
   hm  28. jan.2007   rev 1.1
       modr(x,0) will deliver the result 0

   hm  21. mar 2008    rev 1.2
       use D_trunc for compatibility reasons

   hm  4. apr. 2008    rev 1.3
       added type conversion to avoid warnings under codesys 3.0

   hm  31. oct. 2008   rev 1.4
       changed algorithm to the more common version using floor instead of TRUNC

   hm  10. mar. 2009   rev 1.5
       real constants updated to new systax using dot

   *)
END_FUNCTION

FUNCTION "MUL_ADD" : Real   // FC98, SCL
TITLE = MUL_ADD
{ S7_Optimized_Access := 'FALSE' }
AUTHOR : hugo
FAMILY : MATH
NAME : MUL_ADD
VERSION : 1.1
// this function multiplies an input X with K and adds Offset O to the result.
   VAR_INPUT
      X : Real;
      K : Real;
      O : Real;
   END_VAR
BEGIN


     #MUL_ADD := #X * #K + #O;


   (* revision history
   hm  28. feb 2007
     original version

   hm  11.nov 2007   rev 1.1
     deleted preset values for K and O this makes no sense for a function

   *)
END_FUNCTION

FUNCTION "NEGX" : Real   // FC99, SCL
TITLE = NEGX
{ S7_Optimized_Access := 'FALSE' }
AUTHOR : hugo
FAMILY : MATH
NAME : NEGX
VERSION : 1.0
// This function returns -X
   VAR_INPUT
      X : Real;
   END_VAR
BEGIN


   #NEGX := -#X;

   (* revision history
   hm  26. oct. 2008   rev 1.0
       original version


   *)
END_FUNCTION

FUNCTION "RAD" : Real   // FC100, SCL
TITLE = RAD
{ S7_Optimized_Access := 'FALSE' }
AUTHOR : hugo
FAMILY : MATH
NAME : RAD
VERSION : 1.2
// this function converts Radiant to degrees
// 
// uses: MODR [FC97]
//       FLOOR2 [FC82]
   VAR_INPUT
      deg : Real;
   END_VAR
BEGIN


   #RAD := "MODR"(IN:=0.0174532925199433 * #deg,DIVI:="PI2");

   (*  Enfällt da der Zugriff auf Datenbaustein länger dauert
       RAD := MODR(0.0174532925199433 * DEG, math.PI2);
   *)

   (* revision history
   hm  4. aug 2006     rev 1.0
       original version

   hm  16. oct 2007    rev 1.1
       added modr statement which prohibits rad to become bigger than 2PI

   hm  18. oct 2008    rev 1.2
       using math constants

   *)
END_FUNCTION

FUNCTION "RDM" : Real   // FC101, SCL
TITLE = RDM
{ S7_Optimized_Access := 'FALSE' }
AUTHOR : hugo
FAMILY : MATH
NAME : RDM
VERSION : 1.9
// this function calculates a pseudo random number
// to generate the number it reads the sps timer and calculates a random number between 0 and 1:
// in order to use rdm more then once within one sps cycle it need to be called with different seed numbers LAST.
//  
// uses: T_PLC_MS [FC64]
//       STIME [FB64],IDB_STIME [DB64]
//       BIT_COUNT [FC291]
//       FRACT [FC83]
   VAR_INPUT
      last : Real;
   END_VAR
   VAR_TEMP
      tn : DWord;
      _tn AT tn : Array[0..31] of Bool;
      tc : Int;
   END_VAR
BEGIN


   #tn := "T_PLC_MS"();
   #tc := "BIT_COUNT"(#tn);
   #_tn[7] := #_tn[26];  //tn.31 := tn.2;
   #_tn[6] := #_tn[29];  //tn.30 := tn.5;
   #_tn[5] := #_tn[28];  //tn.29 := tn.4;
   #_tn[4] := #_tn[25];  //tn.28 := tn.1;
   #_tn[3] := #_tn[24];  //tn.27 := tn.0;
   #_tn[2] := #_tn[31];  //tn.26 := tn.7;
   #_tn[1] := #_tn[30];  //tn.25 := tn.6;
   #_tn[0] := #_tn[27];  //tn.24 := tn.3;
   #tn := ROL(IN:=#tn,N:="BIT_COUNT"(#tn)) AND 16#7FFFFFFF OR 16#40000001;  // OR 16#80000001
   #tn := DINT_TO_DWORD(DWORD_TO_DINT(#tn) MOD 71474513 + #tc + 77);
   #RDM := "FRACT"(DINT_TO_REAL(DWORD_TO_DINT(#tn)) / 10000000.0 * ("E"- LIMIT(MN:=0.0,IN:=#last,MX:=1.0)));


   (*
   pt := ADR(temp);
   pt^ := (T_PLC_MS() AND 16#007FFFFF) OR 16#3D000000;
   RDM := fract(modR(temp*e+pi1, PI1-last) + modR(temp*PI1+e + last,e-last));
   *)

   (* revision history
   hm      16. jan 2007        rev 1.0
       original version

   hm      11. nov 2007        rev 1.1
       changed time() into t_plc_ms()

   hm      20. nov 2007        rev 1.2
       changed code of temp calculation to avoid overflow in modr due to resuclt would not fit DINT for high timeer values

   hm      5. jan 2008     rev 1.3
       changed calculation of temp to avoid problem with high values of t_plc_ms

   hm      2. feb 2008     rev 1.4
       changed algorithm to avoind non iec functions and guarantee more randomness

   hm  10. mar. 2008       rev 1.5
       make sure last will be between 0 and 1 to avoid invalid results

   hm  16. mar. 2008       rev 1.6
       added conversion for tc to avoid warnings under codesys 3.0

   hm  18. may. 2008       rev 1.7
       changed constant E to E1

   hm  18. oct. 2008       rev 1.8
       using math constants

   hm  10. mar. 2009       rev 1.9
       real constants updated to new systax using dot

   *)
END_FUNCTION

FUNCTION "RDM2" : Int   // FC102, SCL
TITLE = RDM2
{ S7_Optimized_Access := 'FALSE' }
AUTHOR : hugo
FAMILY : MATH
NAME : RDM2
VERSION : 1.1
// this function calculates an integer pseudo random number
// the random number will be in the range of low <= rdm2 <= high.
// 
// uses: RDM [FC101]
//       T_PLC_MS [FC64] 
//       STIME [FB64],IDB_STIME [DB64] 
//       BIT_COUNT [FC291] 
//       FRACT [FC83]
   VAR_INPUT
      last : Int;
      low : Int;
      high : Int;
   END_VAR
BEGIN


   #RDM2 := REAL_TO_INT(DINT_TO_REAL(TRUNC("RDM"("FRACT"(#last*"PI")) * (#high - #low + 1)) + #low));

   (* revision history
   hm      29. feb 2008        rev 1.0
       original version

   hm      18. oct. 2008       rev 1.1
       using math constants

   *)
END_FUNCTION

FUNCTION "RDMDW" : DWord   // FC103, SCL
TITLE = RDMDW
{ S7_Optimized_Access := 'FALSE' }
AUTHOR : hugo
FAMILY : MATH
NAME : RDMDW
VERSION : 1.2
// this function calculates a DWORD pseudo random number.
// 
// uses: BIT_COUNT [FC291]
//       RDM [FC101]
//       T_PLC_MS [FC64] 
//       STIME [FB64],IDB_STIME [DB64] 
//       FRACT [FC83]
   VAR_INPUT
      last : DWord;
   END_VAR
   VAR_TEMP
      RX : Real;
      "M" : Real;
   END_VAR
BEGIN


   #"M" := "BIT_COUNT"(#last);
   #RX := "RDM"("FRACT"(#"M"*"PI"));
   #RDMDW := SHL(IN:=DINT_TO_DWORD(REAL_TO_DINT(#RX*65535)),N:=16);
   #RX := "RDM"("FRACT"(#"M" * "E"));
   #RDMDW := #RDMDW OR (DINT_TO_DWORD(REAL_TO_DINT(#RX*65535)) AND 16#0000FFFF);

   (* revision history
   hm      14. mar 2008        rev 1.0
       original version

   hm      18. may. 2008       rev 1.1
       changed constant E to E1

   hm      18. oct. 2008       rev 1.2
       using math constants

   *)
END_FUNCTION

FUNCTION "RND" : Real   // FC104, SCL
TITLE = RND
{ S7_Optimized_Access := 'FALSE' }
AUTHOR : hugo
FAMILY : MATH
NAME : RND
VERSION : 1.2
// this function rounds a real down to n digits total.
// round(3.1415,2) = 3.1
// 
// uses: EXPN [FC78]
//       CEIL [FC66]
   VAR_INPUT
      X : Real;
      N : Int;
   END_VAR
   VAR_TEMP
      "M" : Real;
   END_VAR
BEGIN


   IF #X = 0.0 THEN
       #RND := 0.0;
   ELSE
       #"M" := "EXPN"(X:=10.0, N:=#N - "CEIL"((LN(ABS(#X))/LN(10))));
       #RND := DINT_TO_REAL(REAL_TO_DINT(#X * #"M")) / #"M";
   END_IF;


   (* revision history
   hm  11. mar 2008    rev 1.0
       original version

   hm  26. oct. 2008   rev 1.1
       code optimization

   hm  10. mar. 2009   rev 1.2
       real constants updated to new systax using dot

   *)
END_FUNCTION

FUNCTION "ROUND" : Real   // FC105, SCL
TITLE = ROUND
{ S7_Optimized_Access := 'FALSE' }
AUTHOR : hugo
FAMILY : MATH
NAME : ROUND
VERSION : 1.5
// this function rounds a real down to n digits behind the comma.
// round(3.1415,1) = 3.1
   VAR_INPUT
      in : Real;
      N : Int;
   END_VAR
   VAR_TEMP
      X : Real;
   END_VAR
BEGIN


   //x := setup.DECADES[LIMIT(0,n,8)];
   CASE LIMIT(MN:=0, IN:=#N, MX:=8) OF
       1 :           #X:= 10;
       2 :           #X:= 100;
       3 :           #X:= 1000;
       4 :           #X:= 10000;
       5 :           #X:= 100000;
       6 :           #X:= 1000000;
       7 :           #X:= 10000000;
       8 :           #X:= 100000000;
   ELSE: 
       #X:= 1;
   END_CASE ;

   #ROUND := DINT_TO_REAL(REAL_TO_DINT(#in * #X)) / #X;


   (* revision history
   hm  1. sep 2006 rev 1.0
       original version

   hm  2. dec 2007 rev 1.1
       changed code for better performance

   hm  8. jan 2008 rev 1.2
       further improvement in performance

   hm 11. mar. 2008    rev 1.3
       corrected an error with negative numbers
       use real_to_dint instead of trunc

   hm  16. mar 2008    rev 1.4
       added type conversion to avoid warning under codesys 3.0

   hm  25. oct. 2008   rev 1.5
       new code using global constants decades
   *)
END_FUNCTION

FUNCTION "SGN" : Int   // FC106, SCL
TITLE = SGN
{ S7_Optimized_Access := 'FALSE' }
AUTHOR : hugo
FAMILY : MATH
NAME : SGN
VERSION : 1.1
// sgn returns 0 when X = 0 , -1 when X < 1 and +1 when X > 1
   VAR_INPUT
      X : Real;
   END_VAR
BEGIN


     IF #X > 0.0 THEN
       #SGN := 1;
     ELSIF #X < 0.0 THEN
       #SGN := -1;
     ELSE
       #SGN := 0;
     END_IF;

   (* revision histroy
   hm  16. oct 2007  rev 1.0
     original version

   hm  11. nov 2007  rev 1.1
     changed type of function from real to int
   *)
END_FUNCTION

FUNCTION "SIGMOID" : Real   // FC107, SCL
TITLE = SIGMOID
{ S7_Optimized_Access := 'FALSE' }
AUTHOR : hugo
FAMILY : MATH
NAME : SIGMOID
VERSION : 1.2
// this function calculates the sigmoid function
   VAR_INPUT
      X : Real;
   END_VAR
BEGIN


   IF #X > 20.0 THEN
       #SIGMOID := 1.0;
   ELSIF #X < -85.0 THEN
       #SIGMOID := 0.0;
   ELSE
       #SIGMOID := 1.0 / (1.0 + EXP(-#X));
   END_IF;


   (* revision history
   hm  10.12.2007      rev 1.0
       original version

   hm    11. mar. 2008       rev 1.1
       extended range of valid inputs to +inv / -inv

   hm 10. mar. 2009        rev 1.2
       real constants updated to new systax using dot

   *)
END_FUNCTION

FUNCTION "SIGN_I" : Bool   // FC108, SCL
TITLE = SIGN_I
{ S7_Optimized_Access := 'FALSE' }
AUTHOR : hugo
FAMILY : MATH
NAME : SIGN_I
VERSION : 1.3
// this function return true if the integer input is negative
   VAR_INPUT
      IN : DInt;
   END_VAR
BEGIN


   #SIGN_I := #IN < 0;

   (* revision history
   hm 3.3.2007 rev 1.1
       changed method of function for better compatibility to other systems

   hm  1.12.2007   rev 1.2
       changed code to improve performance

   hm  27. oct. 2008   rev 1.3
       changed type of input to dint
   *)
END_FUNCTION

FUNCTION "SIGN_R" : Bool   // FC109, SCL
TITLE = SIGN_R
{ S7_Optimized_Access := 'FALSE' }
AUTHOR : hugo
FAMILY : MATH
NAME : SIGN_R
VERSION : 1.4
// this function return true if the real input is negative
   VAR_INPUT
      in : Real;
   END_VAR
BEGIN


   #SIGN_R := #in < 0.0;


   (* revision history
   hm 19.1.2007    rev 1.1
       changed method of function for better compatibility to other systems

   hm  1.12.2007   rev 1.2
       changed code to improve performance

   hm  14. jun. 2008   rev 1.3
       improved performace

   hm 10. mar. 2009    rev 1.4
       real constants updated to new systax using dot
   *)
END_FUNCTION

FUNCTION "SINC" : Real   // FC110, SCL
TITLE = SINC
{ S7_Optimized_Access := 'FALSE' }
AUTHOR : hugo
FAMILY : MATH
NAME : SINC
VERSION : 1.2
// this function calculates the sinc function.
   VAR_INPUT
      X : Real;
   END_VAR
BEGIN


   IF #X = 0.0 THEN
       #SINC := 1.0;
   ELSE
       #SINC := SIN(#X) / #X;
   END_IF;


   (* revision histroy
   hm  11. mar. 2008   rev 1.0
       original version

   hm  1.12.2007   rev 1.1
       changed code to improove performance

   hm 10. mar. 2009    rev 1.2
       real constants updated to new systax using dot

   *)
END_FUNCTION

FUNCTION "SINH" : Real   // FC111, SCL
TITLE = SINH
{ S7_Optimized_Access := 'FALSE' }
AUTHOR : hugo
FAMILY : MATH
NAME : SINH
VERSION : 1.3
// this function calculates the sin hyperbolicus
   VAR_INPUT
      X : Real;
   END_VAR
BEGIN


   IF ABS(#X) < 2.0E-3 THEN
       #SINH := #X;
   ELSE
       #SINH := (EXP(#X) - EXP(-#X)) * 0.5;
   END_IF;

   (* revision history
   hm  12.1.2007   rev 1.0
       original version

   hm  1.12.2007   rev 1.1
       changed code to improve performance

   hm  5. jan 2008 rev 1.2
       further performance improvement

   hm  11. mar 2008    rev 1.3
       improved accuracy around 0

   *)
END_FUNCTION

FUNCTION "SQRTN" : Real   // FC112, SCL
TITLE = SQRTN
{ S7_Optimized_Access := 'FALSE' }
AUTHOR : hugo
FAMILY : MATH
NAME : SQRTN
VERSION : 1.3
// this function calculates the nth root function of X according to the formula sqrtn = x^(1/n).
   VAR_INPUT
      X : Real;
      N : Int;
   END_VAR
BEGIN


   IF #N > 0 THEN
       #SQRTN := EXP(LN(#X) / INT_TO_REAL(#N));
   ELSE
       #SQRTN := 0.0;
   END_IF;


   (* revision history
   hm      12 jan 2007 rev 1.0
       original version

   hm      2. dec 2007 rev 1.1
       changed code for better performance

   hm      11. mar 2008    rev 1.2
       added result 0 for compatibility reasons

   hm 10. mar. 2009    rev 1.3
       added type conversions for compatibility reasons

   *)
END_FUNCTION

FUNCTION "TANC" : Real   // FC113, SCL
TITLE = TANC
{ S7_Optimized_Access := 'FALSE' }
AUTHOR : hugo
FAMILY : MATH
NAME : TANC
VERSION : 1.1
// this function calculates the tanc function.
   VAR_INPUT
      X : Real;
   END_VAR
BEGIN


   IF #X = 0.0 THEN
       #TANC := 1.0;
   ELSE
       #TANC := TAN(#X) / #X;
   END_IF;


   (* revision histroy
   hm  23. oct. 2008   rev 1.0
       original version

   hm 10. mar. 2009    rev 1.1
       real constants updated to new systax using dot

   *)
END_FUNCTION

FUNCTION "TANH" : Real   // FC114, SCL
TITLE = TANH
{ S7_Optimized_Access := 'FALSE' }
AUTHOR : hugo
FAMILY : MATH
NAME : TANH
VERSION : 1.3
// this function calculates the tangens hyperbolicus
   VAR_INPUT
      X : Real;
   END_VAR
BEGIN


   IF #X > 20.0 THEN
       #TANH := 1.0;
   ELSIF #X < -20.0 THEN
       #TANH := -1.0;
   ELSE
       #TANH := 1.0 - 2.0 / (EXP(2.0 * #X) + 1.0);
   END_IF;


   (* revision hisdtory
   hm      12.1.2007       rev 1.0
       original version

   hm      1.12.2007       rev 1.1
       changed code to improve performance

   hm      10. mar 2008    rev 1.2
       corrected an error in formula
       extended range of valid inputs to +/- INV

   hm 10. mar. 2009    rev 1.3
       real constants updated to new systax using dot

   *)
END_FUNCTION

FUNCTION "WINDOW" : Bool   // FC115, SCL
TITLE = WINDOW
{ S7_Optimized_Access := 'FALSE' }
AUTHOR : hugo
FAMILY : MATH
NAME : WINDOW
VERSION : 1.1
// this checks a signal if the signal is between the upper and lower limit
   VAR_INPUT
      low : Real;
      in : Real;
      high : Real;
   END_VAR
BEGIN


   #WINDOW := #in < #high AND #in > #low;


   (* revision history
   hm  22.1.2007   rev 1.1
       changed the order of inputs to low, in, high

   *)
END_FUNCTION

FUNCTION "WINDOW2" : Bool   // FC116, SCL
TITLE = WINDOW2
{ S7_Optimized_Access := 'FALSE' }
AUTHOR : hugo
FAMILY : MATH
NAME : WINDOW2
VERSION : 1.0
// this checks a signal if the signal is between the upper and lower limit including the two limits
   VAR_INPUT
      low : Real;
      in : Real;
      high : Real;
   END_VAR
BEGIN


   #WINDOW2 := #in <= #high AND #in >= #low;


   (* revision history
   hm  31.10.2007  rev 1.0
     original version

   *)
END_FUNCTION

FUNCTION "BIT_COUNT" : Int   // FC291, SCL
TITLE = BIT_COUNT
{ S7_Optimized_Access := 'FALSE' }
AUTHOR : hugo
FAMILY : GATE
NAME : BITCT
VERSION : 1.1
// BIT_COUNT counts the amount True of bits in a dword.
// for exabple: bit_count(3) returns 2 because two bits (bits 0 and 1) are true and all others are false.
   VAR_INPUT
      IN : DWord;
   END_VAR
   VAR_TEMP
      temp : DWord;
      attemp AT temp : Array[0..31] of Bool;
   END_VAR
BEGIN


     #BIT_COUNT := 0;
     #temp := #IN;

     WHILE DWORD_TO_DINT(#temp) <> 0 DO
       IF #attemp[24] THEN #BIT_COUNT := #BIT_COUNT +1; END_IF;
       #temp := SHR(IN:=#temp,N:=1);
     END_WHILE;

   (* revision history
   5.7.2007  rev 1.0    original version

   10.9.2007  rev 1.1    hm
     changed algorithm for better performace
     the execution time has reduced by a factor of 5
     deleted unused variable temp
   *)
END_FUNCTION

FUNCTION "LAMBERT_W" : Real   // FC414, SCL
TITLE = LAMBERT_W
{ S7_Optimized_Access := 'FALSE' }
AUTHOR : hugo
FAMILY : MATH
NAME : LAMBERT
VERSION : 1.1
// this function calculates the lambert_w function.
   VAR_INPUT
      X : Real;
   END_VAR
   VAR_TEMP
      w : Real;
      i : Int;
      we : Real;
      w1e : Real;
      last : DWord;
      ewx : Real;
   END_VAR
BEGIN


   (* check for valid input and return -1000 if too low *)
   IF #X < -0.367879441171442 THEN
       #LAMBERT_W := -1000.0;
       RETURN;
   (* return 0 if x = 0 *)
   ELSIF #X = 0.0 THEN
       RETURN;
   (* first an estimate is calculated *)
   ELSIF #X <= 500.0 THEN
       #w := LN(#X + 1.0);
       #w := 0.665 * (1.0 + 0.0195 * #w) * #w + 0.04;
   ELSE
       #w := LN(#X - 4.0) - (1.0 - 1.0/LN(#X)) * LN(LN(#X));
   END_IF;
   (* use estimate to calculate exact result *)
   FOR #i := 0 TO 5 DO
       #ewx := EXP(#w);
       #we := #w * #ewx - #X;
       #w1e := (#w + 1.0) * #ewx;
       #last := REAL_TO_DWORD(#w) AND 16#FFFF_FFFC;
       #w := #w - (#we / (#w1e - (#w+2.0) * #we / (2.0 * #w + 2.0)));
       IF (REAL_TO_DWORD(#w) AND 16#FFFF_FFFC) = #last THEN EXIT; END_IF;
   END_FOR;
   #LAMBERT_W := #w;


   (* revision hisdtory
   hm  26. oct. 2008   rev 1.0
       original version

   hm  10. mar. 2009   rev 1.1
       real constants updated to new systax using dot

   *)
END_FUNCTION

FUNCTION "REAL_TO_FRAC" : "FRACTION"   // FC427, SCL
TITLE = REAL_TO_FRAC
{ S7_Optimized_Access := 'FALSE' }
AUTHOR : alex
FAMILY : MATH
NAME : R2FRAC
VERSION : 1.0
// this function calculates the closest fraction for a real number
// 
// uses: FRACTION [UDT19]
   VAR_INPUT
      X : Real;
      N : Int;
   END_VAR
   VAR_TEMP
      temp : DInt;
      sign : Bool;
      X_gerundet : DInt;
      X_ohne_Nachkomma : Real;
      Numerator : DInt;
      Denominator : DInt;
      Numerator_old : DInt;
      Denominator_old : DInt;
      tX : Real;
      tREAL_TO_FRAC : "FRACTION";
   END_VAR
BEGIN


   #Numerator := 1; (* Initialwert Zaehler  *)
   #Denominator := 0; (* Initialwert Nenner *)
   #Numerator_old := 0; (* Initialwert Zaehler der letzten Berechnung  *)
   #Denominator_old := 1; (* Initialwert Zaehler der letzten Berechnung   *)
   #tX := #X;

   (*
   numerator := 1;                     (* Zaehler Initialwert *)
   denominator := 0;                   (* Nenner  Initialwert *)
   numerator_old := 0;
   denominator_old :=1;
   *)

   IF #tX < 0.0 THEN
     #sign := TRUE;               (* Vorzeichen merken *)
     #tX := ABS(#tX);              (* Absolutwert berechnen *)
   END_IF;

   (*
   sign := SIGN_R(X);                    
   X := ABS(X);                      
   *)

   REPEAT
     #X_gerundet := REAL_TO_DINT(#tX);

     (* Zaehler berechnen *)
     #temp := #Numerator * #X_gerundet + #Numerator_old;   (* Zaehler um Vorkammawert erweitern *)
     #Numerator_old := #Numerator;             (* Zaehler der letzten Berechnung speichern *)
     #Numerator := #temp;                  (* Zaehler dieser Berechnung speichern *)

     (* Nenner berechnen *)
     #temp := #Denominator * #X_gerundet + #Denominator_old; (* Nenner um Vorkammawert erweitern *)
     #Denominator_old := #Denominator;           (* Nenner der letzten Berechnung speichern *)
     #Denominator := #temp;                (* Nenner dieser Berechnung speichern *)

     (* Restwert berechnen *)
     #X_ohne_Nachkomma := DINT_TO_REAL(#X_gerundet);
     IF #tX = #X_ohne_Nachkomma THEN            (* Bruch geht ohne Rest auf *)
       IF ABS(#Denominator) <= #N THEN         (* kein Rundungsfehler *)
         #Numerator_old := #Numerator;         (* Numerator_old wird von Funktion zurückgegeben *)
         #Denominator_old := #Denominator;       (* Denominator_old wird von Funktion zurückgegeben *)
       END_IF;
       EXIT;                     (* keine weitere Berechnung notwendig *)
     ELSE
       #tX := 1.0 / (#tX - #X_ohne_Nachkomma);        (* Kehrwert vom Rest -> Neuer Bruch *)
     END_IF;

   UNTIL
     ( ABS(#Denominator) > #N )
   END_REPEAT;

   (* correct sign if X was negative *)
   IF #sign THEN
     #tREAL_TO_FRAC.NUMERATOR := -1 * ABS(DINT_TO_INT(#Numerator_old));
   ELSE
     #tREAL_TO_FRAC.NUMERATOR :=  ABS(DINT_TO_INT(#Numerator_old));
   END_IF;

   #tREAL_TO_FRAC.DENOMINATOR := ABS(DINT_TO_INT(#Denominator_old));

   #REAL_TO_FRAC := #tREAL_TO_FRAC;


   (* revision history
   hm    19. jan. 2011 rev 1.0
     original version

   ad    06. apr. 2011 rev 1.1
     optimized code
   *)
END_FUNCTION

FUNCTION "GCD" : Int   // FC431, SCL
TITLE = GCD
{ S7_Optimized_Access := 'FALSE' }
AUTHOR : hugo
FAMILY : MATH
NAME : GCD
VERSION : 1.0
// this function calculates the gretaest common divisor of two numbers A and B
   VAR_INPUT
      "A" : DInt;
      "B" : DInt;
   END_VAR
   VAR_TEMP
      t : DInt;
      tA : DInt;
      _A AT tA : Array[0..31] of Bool;
      tB : DInt;
      _B AT tB : Array[0..31] of Bool;
   END_VAR
BEGIN


   #tA := #"A";
   #tB := #"B";

   IF #tA = 0 THEN
     #GCD := DINT_TO_INT(ABS(#tB));
   ELSIF #tB = 0 THEN
     #GCD := DINT_TO_INT(ABS(#tA));
   ELSE
     #tA := ABS(#tA);
     #tB := ABS(#tB);
     #GCD := 1;
     WHILE NOT(#_A[24] OR #_B[24]) DO
       #tA := DWORD_TO_DINT(SHR(IN:=DINT_TO_DWORD(#tA),N:=1));
       #tB := DWORD_TO_DINT(SHR(IN:=DINT_TO_DWORD(#tB),N:=1));
       #GCD := WORD_TO_INT(SHL(IN:=INT_TO_WORD(#GCD),N:=1));
     END_WHILE;
     WHILE #tA > 0 DO
       IF NOT(#_A[24]) THEN #tA := DWORD_TO_DINT(SHR(IN:=DINT_TO_DWORD(#tA),N:=1));
       ELSIF NOT(#_B[24]) THEN #tB := DWORD_TO_DINT(SHR(IN:=DINT_TO_DWORD(#tB),N:=1));
       ELSE
         #t:= DWORD_TO_DINT(SHR(IN:=DINT_TO_DWORD(ABS(#tA-#tB)),N:=1));
         IF #tA < #tB THEN #tB := #t; ELSE #tA := #t; END_IF;
       END_IF;
     END_WHILE;
     #GCD := #GCD * DINT_TO_INT(#tB);
   END_IF;


   (* revision history
   hm  19. jan. 2011 rev 1.0
     original version

   *)
END_FUNCTION

// ===== PLC "Mathematical Array"  Unspecific CPU S7 300 =====

VAR_GLOBAL CONSTANT   // PLC tag table "STEP7 classic symbols"
   "debug" : Bool := FALSE;
   "N" : Int := 0;
   "offset" : Int := 0;
   "E" : Real := 2.71828182845904523536028747135266249;   // Eulersche Konstante
   "PI" : Real := 3.14159265358979323846264338327950288;
   "offset_1" : DWord := 0;
END_VAR

DATA_BLOCK "IDB_STIME"   // DB64
{ S7_Optimized_Access := 'FALSE' }
AUTHOR : dalbi
FAMILY : MEASURE
VERSION : 0.0
// stored: InstanceOfName STIME
"STIME"
BEGIN
END_DATA_BLOCK

FUNCTION_BLOCK "_ARRAY_ABS"   // FB5, SCL
TITLE = _ARRAY_ABS
{ S7_Optimized_Access := 'FALSE' }
AUTHOR : hugo
FAMILY : ARFUNCT
NAME : AR_ABS
VERSION : 1.0
// this function will calculate the absolute value of each element of the array and stroe the result instead of the element.
// Array[i] := ABS(ARRAY[i]).
// the function needs to be called:    array_avg(adr("array"),sizeof("array"));
// because this function works with pointers its very time efficient and it needs no extra memory.
   VAR_INPUT
      pt : Pointer;
      _pt AT pt : Struct
         DBNr : Word;
         Adr : DWord;
      END_STRUCT;
      size : Int;
   END_VAR
   VAR_OUTPUT
      _ABS : Bool;
   END_VAR
   VAR_TEMP
      i : Int;
      stop : Int;
      Adr : Int;
      DB_LENGTH : Word;
      WRITE_PROT : Bool;
      rTEST_DB : Int;
   END_VAR
BEGIN


   #_ABS := FALSE;

   (* test data block *)
   #rTEST_DB := TEST_DB(DB_NUMBER := #_pt.DBNr ,DB_LENGTH => #DB_LENGTH ,WRITE_PROT => #WRITE_PROT);
   (* End if TEST_DB <> 0 = Error *)
   IF #rTEST_DB <> 0 THEN RETURN; END_IF;
   (* End if data block to short *) 
   IF WORD_TO_INT(#DB_LENGTH)/4 < #size THEN RETURN; END_IF;
   (* calculate adress for first data *)  
   #Adr := DWORD_TO_INT(SHR(IN:=SHL(IN:=#_pt.Adr,N:=8),N:=11));

   (* code *)
   #stop := #size - 1;   //stop := SHR(size,2)-1;
   FOR #i := 0 TO #stop DO
       WORD_TO_BLOCK_DB(#_pt.DBNr).DD(#Adr+#i*4) := REAL_TO_DWORD(ABS(DWORD_TO_REAL(WORD_TO_BLOCK_DB(#_pt.DBNr).DD(#Adr+#i*4))));
   END_FOR;

   #_ABS := TRUE;


   (* revision history
   hm  2. apr 2008     rev 1.0
       original version

   *)
END_FUNCTION_BLOCK

FUNCTION_BLOCK "_ARRAY_ADD"   // FB6, SCL
TITLE = _ARRAY_ADD
{ S7_Optimized_Access := 'FALSE' }
AUTHOR : hugo
FAMILY : ARFUNCT
NAME : AR_ADD
VERSION : 1.0
// this function will add an offset X to each element of the array and stroe the result instead of the element.
// Array[i] := ARRAY[i] + X.
// the function needs to be called:    array_avg(adr("array"),sizeof("array"));
// because this function works with pointers its very time efficient and it needs no extra memory.
   VAR_INPUT
      pt : Pointer;
      _pt AT pt : Struct
         DBNr : Word;
         Adr : DWord;
      END_STRUCT;
      size : Int;
      X : Real;
   END_VAR
   VAR_OUTPUT
      _ADD : Bool;
   END_VAR
   VAR_TEMP
      i : Int;
      stop : Int;
      Adr : Int;
      DB_LENGTH : Word;
      WRITE_PROT : Bool;
      rTEST_DB : Int;
   END_VAR
BEGIN


   #_ADD := FALSE;

   (* test data block *)
   #rTEST_DB := TEST_DB(DB_NUMBER := #_pt.DBNr ,DB_LENGTH => #DB_LENGTH ,WRITE_PROT => #WRITE_PROT);
   (* End if TEST_DB <> 0 = Error *)
   IF #rTEST_DB <> 0 THEN RETURN; END_IF;
   (* End if data block to short *) 
   IF WORD_TO_INT(#DB_LENGTH)/4 < #size THEN RETURN; END_IF;
   (* calculate adress for first data *)  
   #Adr := DWORD_TO_INT(SHR(IN:=SHL(IN:=#_pt.Adr,N:=8),N:=11));

   (* code *)
   #stop := #size - 1;   //stop := SHR(size,2)-1;
   FOR #i := 0 TO #stop DO
       WORD_TO_BLOCK_DB(#_pt.DBNr).DD(#Adr+#i*4) := REAL_TO_DWORD(DWORD_TO_REAL(WORD_TO_BLOCK_DB(#_pt.DBNr).DD(#Adr+#i*4)) + #X);
   END_FOR;
   #_ADD := TRUE;


   (* revision history
   hm  2. apr 2008     rev 1.0
       original version

   *)
END_FUNCTION_BLOCK

FUNCTION_BLOCK "_ARRAY_INIT"   // FB7, SCL
TITLE = _ARRAY_INIT
{ S7_Optimized_Access := 'FALSE' }
AUTHOR : hugo
FAMILY : ARFUNCT
NAME : AR_INIT
VERSION : 1.3
// this function will initialize a given array with a value init.
// the function needs to be called:    _array_init(adr("array"),sizeof("array"));
// this function will manipulate a given array.
// the function manipulates the original array, it rerturnes true when finished.
// because this function works with pointers its very time efficient and it needs no extra memory.
   VAR_INPUT
      pt : Pointer;
      _pt AT pt : Struct
         DBNr : Word;
         Adr : DWord;
      END_STRUCT;
      size : Int;
      init : Real;
   END_VAR
   VAR_OUTPUT
      _init : Bool;
   END_VAR
   VAR_TEMP
      i : Int;
      Adr : Int;
      DB_LENGTH : Word;
      WRITE_PROT : Bool;
      rTEST_DB : Int;
   END_VAR
BEGIN


     #_init := FALSE;

     (* Datenbaustein Testen *)
     #rTEST_DB := TEST_DB(DB_NUMBER := #_pt.DBNr // IN: WORD
                        ,DB_LENGTH => #DB_LENGTH // OUT: WORD
                        ,WRITE_PROT => #WRITE_PROT // OUT: BOOL
                        ); // INT
     (* Ende wenn Test-DB <> 0 = Fehler *)
     IF #rTEST_DB <> 0 THEN RETURN; END_IF;
     (* Ende wenn DB zu klein *) 
     IF WORD_TO_INT(#DB_LENGTH)/4 < #size THEN RETURN; END_IF;

     #Adr := DWORD_TO_INT(SHR(IN:=SHL(IN:=#_pt.Adr,N:=8),N:=11));

     (* Berechnung *)
     FOR #i := 0 TO #size-1 DO
         WORD_TO_BLOCK_DB(#_pt.DBNr).DD(#Adr+#i*4) := REAL_TO_DWORD(#init);    
     END_FOR;
     #_init := TRUE;

   (* revision History

   hm 6.1.2007     rev 1.1
       change type of function to bool
       added  array_init := true to set output true.

   hm  14.11.2007  rev 1.2
       changed stop calculation to be more efficient

   hm  16.3. 2008      rev 1.3
       changed type of input size to uint
   *)
END_FUNCTION_BLOCK

FUNCTION_BLOCK "_ARRAY_MEDIAN"   // FB8, SCL
TITLE = _ARRAY_MEDIAN
{ S7_Optimized_Access := 'FALSE' }
AUTHOR : hugo
FAMILY : ARFUNCT
NAME : AR_MEDI
VERSION : 1.5
// this function will calculate the median of a given array.
// in order to do so the ariginal array is sorted and stays sorted after the function finishes
// the function needs to be called:    _array_median(adr("array"),sizeof("array"));
// this function will manipulate a given array.
// the function will return the median of the original array.
// for example [12,0,4,7,1] the median is 4 and the array after the function is called is [0,1,4,7,12]
// because this function works with pointers its very time efficient and it needs no extra memory.
// 
// uses: EVEN [FC76]
//       _ARRAY_SORT [FB11]
   VAR_INPUT
      pt : Pointer;
      at_pt AT pt : Struct
         DBNr : Word;
         Adr : DWord;
      END_STRUCT;
      size : Int;
   END_VAR
   VAR_OUTPUT
      median : Real;
   END_VAR
   VAR
      sort : "_ARRAY_SORT";
   END_VAR
   VAR_TEMP
      i : Int;
      "m" : Int;
      temp : Real;
      stop : Int;
      Adr : Int;
      DB_LENGTH : Word;
      WRITE_PROT : Bool;
      rTEST_DB : Int;
   END_VAR
BEGIN


     (* Datenbaustein Testen *)
     #rTEST_DB := TEST_DB(DB_NUMBER := #at_pt.DBNr // IN: WORD
                        ,DB_LENGTH => #DB_LENGTH // OUT: WORD
                        ,WRITE_PROT => #WRITE_PROT // OUT: BOOL
                        ); // INT
     (* Ende wenn Test-DB <> 0 = Fehler *)
     IF #rTEST_DB <> 0 THEN RETURN; END_IF;
     (* Ende wenn DB zu klein *) 
     IF WORD_TO_INT(#DB_LENGTH)/4 < #size THEN RETURN; END_IF;

     #Adr := DWORD_TO_INT(SHR(IN:=SHL(IN:=#at_pt.Adr,N:=8),N:=11));

     #sort(PT:=#pt,SIZE:=#size);
     #stop := #size-1;
     IF "EVEN"(#stop) THEN
       #median := DWORD_TO_REAL(WORD_TO_BLOCK_DB(#at_pt.DBNr).DD(#Adr+(#stop/2)*4));
     ELSE
       #i := WORD_TO_INT(SHR(IN:=INT_TO_WORD(#stop),N:=1));
       #median := (DWORD_TO_REAL(WORD_TO_BLOCK_DB(#at_pt.DBNr).DD(#Adr+#i*4)) + DWORD_TO_REAL(WORD_TO_BLOCK_DB(#at_pt.DBNr).DD(#Adr+(#i+1)*4)))/2;
     END_IF;

   (* old code
   stop := (size - SIZEOF(pt)) / SIZEOF(pt);
   FOR i := 0 TO stop - 1 DO
       FOR m := i + 1 TO stop DO
           IF pt^[i] > pt^[m] THEN
               temp := pt^[i];
               pt^[i] := pt^[m];
               pt^[m] := temp;
           END_IF;
       END_FOR;
   END_FOR;
   IF even(stop) THEN
       _array_median := pt^[stop/2];
   ELSE
       i := stop/2;
       _array_median := (pt^[i] + pt^[i+1])/2;
   END_IF;
   *)
   (* revision history
   hm  3.3.2007        rev 1.1
       corrected an error, changed the statement line 14    i := TRUNC(stop/2); to i := stop/2;

   hm      22. sep 2007    rev 1.2
       changed algorithm to use _array_soft for performance reasons

   hm      8. oct 2007     rev 1.3
       deleted unused variables m and temp

   hm      14. nov 2007    rev 1.4
       corrected a problem with size calculation

   hm      16.3. 2008      rev 1.5
       changed type of input size to uint
       performance improvements
   *)
END_FUNCTION_BLOCK

FUNCTION_BLOCK "_ARRAY_MUL"   // FB9, SCL
TITLE = _ARRAY_MUL
{ S7_Optimized_Access := 'FALSE' }
AUTHOR : hugo
FAMILY : ARFUNCT
NAME : AR_MUL
VERSION : 1.0
// this function will multiply each element of the array and stroe the result instead of the element.
// Array[i] := ARRAY[i] * X.
// the function needs to be called:    array_avg(adr("array"),sizeof("array"));
// because this function works with pointers its very time efficient and it needs no extra memory.
   VAR_INPUT
      pt : Pointer;
      _pt AT pt : Struct
         DBNr : Word;
         Adr : DWord;
      END_STRUCT;
      size : Int;
      X : Real;
   END_VAR
   VAR_OUTPUT
      _MUL : Bool;
   END_VAR
   VAR_TEMP
      i : Int;
      stop : Int;
      Adr : Int;
      DB_LENGTH : Word;
      WRITE_PROT : Bool;
      rTEST_DB : Int;
   END_VAR
BEGIN


   #_MUL := FALSE;

   (* test data block *)
   #rTEST_DB := TEST_DB(DB_NUMBER := #_pt.DBNr ,DB_LENGTH => #DB_LENGTH ,WRITE_PROT => #WRITE_PROT);
   (* End if TEST_DB <> 0 = Error *)
   IF #rTEST_DB <> 0 THEN RETURN; END_IF;
   (* End if data block to short *) 
   IF WORD_TO_INT(#DB_LENGTH)/4 < #size THEN RETURN; END_IF;
   (* calculate adress for first data *)  
   #Adr := DWORD_TO_INT(SHR(IN:=SHL(IN:=#_pt.Adr,N:=8),N:=11));

   (* code *)
   #stop := #size - 1;   //stop := SHR(size,2)-1;
   FOR #i := 0 TO #stop DO
       WORD_TO_BLOCK_DB(#_pt.DBNr).DD(#Adr+#i*4) := REAL_TO_DWORD(DWORD_TO_REAL(WORD_TO_BLOCK_DB(#_pt.DBNr).DD(#Adr+#i*4)) * #X);
   END_FOR;
   #_MUL := TRUE;


   (* revision history
   hm  2. apr 2008     rev 1.0
       original version

   *)
END_FUNCTION_BLOCK

FUNCTION_BLOCK "_ARRAY_SHUFFLE"   // FB10, SCL
TITLE = _ARRAY_SHUFFLE
{ S7_Optimized_Access := 'FALSE' }
AUTHOR : kurt
FAMILY : ARFUNCT
NAME : AR_SHUFF
VERSION : 1.2
// this function will randomly shuffle the elements of an array
// 
// uses: RDM2 [FC102]
//       RDM [FC101] 
//       T_PLC_MS [FC64]
//       STIME [FB64],IDB_STIME [DB64]
//       BIT_COUNT [FC291]
//       FRACT [FC83]
   VAR_INPUT
      pt : Pointer;
      _pt AT pt : Struct
         DBNr : Word;
         Adr : DWord;
      END_STRUCT;
      size : Int;
   END_VAR
   VAR_OUTPUT
      ARRAY_SHUFFLE : Bool;
   END_VAR
   VAR_TEMP
      temp : Real;
      pos : Int;
      i : Int;
      stop : Int;
      Adr : Int;
      DB_LENGTH : Word;
      WRITE_PROT : Bool;
      rTEST_DB : Int;
   END_VAR
BEGIN


   #ARRAY_SHUFFLE := FALSE;

   (* Datenbaustein Testen *)
   #rTEST_DB := TEST_DB(DB_NUMBER := #_pt.DBNr // IN: WORD
                      ,DB_LENGTH => #DB_LENGTH // OUT: WORD
                      ,WRITE_PROT => #WRITE_PROT // OUT: BOOL
                      ); // INT
   (* Ende wenn Test-DB <> 0 = Fehler *)
   IF #rTEST_DB <> 0 THEN RETURN; END_IF;
   (* Ende wenn DB zu klein *) 
   IF WORD_TO_INT(#DB_LENGTH)/4 < #size THEN RETURN; END_IF;

   #Adr := DWORD_TO_INT(SHR(IN:=SHL(IN:=#_pt.Adr,N:=8),N:=11));

   #stop := #size - 1;//WORD_TO_INT(SHR(IN:=INT_TO_WORD(size),N:=2))-1;
   FOR #i := 0 TO #stop DO
           #pos := "RDM2"(last:=#i+#pos,low:=0,high:=#stop);
           (* swap elements *)
           #temp := DWORD_TO_REAL(WORD_TO_BLOCK_DB(#_pt.DBNr).DD(#Adr+#i*4));
           WORD_TO_BLOCK_DB(#_pt.DBNr).DD(#Adr+#i*4) := WORD_TO_BLOCK_DB(#_pt.DBNr).DD(#Adr+#pos*4);
           WORD_TO_BLOCK_DB(#_pt.DBNr).DD(#Adr+#pos*4) := REAL_TO_DWORD(#temp);
   END_FOR;
   #ARRAY_SHUFFLE := TRUE;


   (* revision History
   hm  4. mar 2008 rev 1.0
       original version

   hm  16. mar. 2008   rev 1.1
       changed type of input size to uint

   hm  30. mar. 2008   rev 1.2
       changed last in rdm2 fromm pos to i + pos to allow for more randomness

   *)
END_FUNCTION_BLOCK

FUNCTION_BLOCK "_ARRAY_SORT"   // FB11, SCL
TITLE = _ARRAY_SORT
{ S7_Optimized_Access := 'FALSE' }
AUTHOR : Alex
FAMILY : ARFUNCT
NAME : AR_SORT
VERSION : 2.0
// this function will sort a given array.
// the function needs to be called:  _array_sort(adr("array"),sizeof("array"));
// this function will manipulate a given array.
// the function will not return anything except true, it will instead manipulate the original array.
// because this function works with pointers its very time efficient and it needs no extra memory.
   VAR_INPUT
      PT : Pointer;
      _PT AT PT : Struct
         DBNr : Word;
         Adr : DWord;
      END_STRUCT;
      SIZE : Int;
   END_VAR
   VAR_OUTPUT
      SORT : Bool;
   END_VAR
   VAR
      stack : Array[1..32] of Int;
   END_VAR
   VAR_TEMP
      stack_count : Int;
      links : Int;
      rechts : Int;
      pivot : Real;
      i : Int;
      j : Int;
      ende_innen : Bool;
      ende_aussen : Bool;
      tmp : Real;
      Adr : Int;
      DB_LENGTH : Word;
      WRITE_PROT : Bool;
      rTEST_DB : Int;
   END_VAR
BEGIN


   #SORT := FALSE;

   (* Datenbaustein Testen *)
   #rTEST_DB := TEST_DB(DB_NUMBER := #_PT.DBNr // IN: WORD
                      ,DB_LENGTH => #DB_LENGTH // OUT: WORD
                      ,WRITE_PROT => #WRITE_PROT // OUT: BOOL
                      ); // INT
   (* Ende wenn Test-DB <> 0 = Fehler *)
   IF #rTEST_DB <> 0 THEN RETURN; END_IF;
   (* Ende wenn DB zu klein *) 
   IF WORD_TO_INT(#DB_LENGTH)/4 < #SIZE THEN RETURN; END_IF;

   #Adr := DWORD_TO_INT(SHR(IN:=SHL(IN:=#_PT.Adr,N:=8),N:=11))-4;

   (* Startwerte zur Arraygröße *)
   #links := 1;         (* Anfangselement des Arrays *)
   #rechts := WORD_TO_INT(SHR(IN:=INT_TO_WORD(#SIZE),N:=2));    (* Endelement des Arrays *)
   #stack_count := 1;     (* Laufvariable Stack *)

   WHILE NOT #ende_aussen DO            (* äußere Schleife *)
     IF #links < #rechts THEN
       #pivot := DWORD_TO_REAL(WORD_TO_BLOCK_DB(#_PT.DBNr).DD((#Adr+WORD_TO_INT(SHR(IN:=INT_TO_WORD(#rechts+#links),N:=1)))*4));      (* Wert des mittleren Elements als Pivot-Wert *)
       #i := #links -1;
       #j := #rechts +1;

       (* innere Schleife, teile Feld *)
       #ende_innen := FALSE;
       REPEAT

         (* steigende Reihenfolge *)
         REPEAT  #i := #i+1; UNTIL (DWORD_TO_REAL(WORD_TO_BLOCK_DB(#_PT.DBNr).DD((#Adr+#i)*4)) >= #pivot) OR NOT (#i < #rechts) END_REPEAT;
         REPEAT  #j := #j-1; UNTIL (DWORD_TO_REAL(WORD_TO_BLOCK_DB(#_PT.DBNr).DD((#Adr+#j)*4)) <= #pivot) OR NOT (#j > #links)  END_REPEAT;


         (*sinkende Reihenfolge *)
   (*      REPEAT  i := i+1; UNTIL (PT^[i] <= pivot) OR NOT (i < rechts) END_REPEAT  *)
   (*      REPEAT  j := j-1; UNTIL (PT^[j] >= pivot) OR NOT (j > links)  END_REPEAT  *)

         IF #i >= #j THEN
           #ende_innen := TRUE;
         ELSE
              #tmp := DWORD_TO_REAL(WORD_TO_BLOCK_DB(#_PT.DBNr).DD((#Adr+#j)*4));
           WORD_TO_BLOCK_DB(#_PT.DBNr).DD((#Adr+#j)*4) := WORD_TO_BLOCK_DB(#_PT.DBNr).DD((#Adr+#i)*4);
           WORD_TO_BLOCK_DB(#_PT.DBNr).DD((#Adr+#i)*4) := REAL_TO_DWORD(#tmp);
         END_IF;

       UNTIL #ende_innen END_REPEAT;

       (* Push stack *)
       #stack[#stack_count] := #rechts;   (* rechten Teil später sortieren *)
       IF #stack_count < 32 THEN
         #stack_count := #stack_count +1;
       ELSE
         #ende_aussen := TRUE;
         #SORT := FALSE;         (* Fehler: Stack zu klein *)
       END_IF;

       (* linken Teil sortiern *)
       #rechts := MAX(IN1:=#links,IN2:=#i-1);

     ELSE

       IF #stack_count = 1 THEN
         #ende_aussen := TRUE;
       ELSE

         #links := #rechts+1;

         (* pop stack *)
         #stack_count := #stack_count -1;    (* jetzt rechten Teil sortierne *)
         #rechts:= #stack[#stack_count];
       END_IF;

     END_IF;

   END_WHILE;

   #SORT := TRUE;        (* Sortierung beendet *)


   (* algorithm used before rev 2.0

   size := SHR(size,2);
   size2 := UINT_TO_INT(SHR(size,1));
   FOR i := SIZE2  TO 1 BY -1 DO
     j:=i;
       WHILE j <= SIZE2 DO
         stop := j * 2 + 1;
           IF stop > UINT_TO_INT(SIZE) THEN stop := stop - 1;
           ELSIF pt^[stop-1] > pt^[stop] THEN stop := stop - 1;
       END_IF;
           IF pt^[j] < pt^[stop] THEN
             temp := pt^[j];
               pt^[j] := pt^[stop];
               pt^[stop] := temp;
           END_IF;
           j := stop;
       END_WHILE;
   END_FOR;

   *)

   (* heapsort
   FOR heapsize := UINT_TO_INT(size) TO 1 BY -1 DO
     popmax := pt^[1];
     pt^[1] := pt^[heapsize];
       i := 1;
     hs2 := SHR(heapsize,1);
     WHILE i <= hs2 DO
           stop := i * 2 + 1;  
             IF stop > heapsize THEN stop := stop - 1;
             ELSIF pt^[stop-1] > pt^[stop] THEN stop := stop - 1;
       END_IF;
             IF pt^[i] < pt^[stop] THEN
                   temp := pt^[i];
                   pt^[i] := pt^[stop];
                   pt^[stop] := temp;
             END_IF;
             i := stop;
         END_WHILE;
     pt^[heapsize] := popmax;
   END_FOR;

   _ARRAY_SORT2 := TRUE;
   *)

   (* old algorithm bubble sort used before rev 1.2
   stop := (size - SIZEOF(pt)) / SIZEOF(pt);
   FOR i := 0 TO stop - 1 DO
     FOR m := i + 1 TO stop DO
       IF pt^[i] > pt^[m] THEN
         temp := pt^[i];
         pt^[i] := pt^[m];
         pt^[m] := temp;
       END_IF;
     END_FOR;
   END_FOR;
   _array_sort := TRUE;

   *)


   (* revision history

   hm  6.1.2007  rev 1.1
     changed return value to true

   hm  22. sep 2007  rev 1.2
     changed sorting algorithm to heap sort for performance reasons

   hm  14. nov 2007  rev 1.3
     changed calculation of stop to be more efficient

   hm  15 dec 2007 rev 1.4
     added function return true

   hm  5. jan 2008   rev 1.5
     improved performance

   hm  16. mar. 2008 rev 1.6
     changed type of input size to uint

   hm  28. mar. 2008 rev 1.7
     changed input f to pt

   hm  19. jan. 2011 rev 2.0
     new faster algorithm using qucksort (Alexander Drikitis)

   *)
END_FUNCTION_BLOCK

FUNCTION_BLOCK "ARRAY_AVG"   // FB12, SCL
TITLE = ARRAY_AVG
{ S7_Optimized_Access := 'FALSE' }
AUTHOR : hugo
FAMILY : ARFUNCT
NAME : AR_AVG
VERSION : 1.3
// this function will calculate the average of a given array.
// the function needs to be called:  array_avg(adr("array"),sizeof("array"));
// because this function works with pointers its very time efficient and it needs no extra memory.
   VAR_INPUT
      pt : Pointer;
      _pt AT pt : Struct
         DBNr : Word;
         Adr : DWord;
      END_STRUCT;
      size : Int;
   END_VAR
   VAR_OUTPUT
      avg : Real;
   END_VAR
   VAR_TEMP
      i : Int;
      stop : Int;
      Adr : Int;
      DB_LENGTH : Word;
      WRITE_PROT : Bool;
      rTEST_DB : Int;
   END_VAR
BEGIN


   (* Datenbaustein Testen *)
   #rTEST_DB := TEST_DB(DB_NUMBER := #_pt.DBNr, DB_LENGTH => #DB_LENGTH, WRITE_PROT => #WRITE_PROT);
   (* Ende wenn Test-DB <> 0 = Fehler *)
   IF #rTEST_DB <> 0 THEN RETURN; END_IF;
   (* Ende wenn DB zu klein *) 
   IF WORD_TO_INT(#DB_LENGTH)/4 < #size THEN RETURN; END_IF;

   #Adr := DWORD_TO_INT(SHR(IN:=SHL(IN:=#_pt.Adr,N:=8),N:=11));

   #stop := #size-1;
   #avg := DWORD_TO_REAL(WORD_TO_BLOCK_DB(#_pt.DBNr).DD(#Adr+0));
   FOR #i := 1 TO #stop DO
       #avg := #avg + DWORD_TO_REAL(WORD_TO_BLOCK_DB(#_pt.DBNr).DD(#Adr+#i*4));
   END_FOR;
   #avg := #avg / INT_TO_REAL(#stop + 1);


   (* revision history
   hm  2. oct 2007     rev 1.0
       original version

   hm  12. dec 2007    rev 1.1
       chaged code for better performance

   hm  16. mar. 2008   rev 1.2
       changed input size to uint

   hm  10. mar. 2009   rev 1.3
       added type conversion for compatibility reasons
   *)
END_FUNCTION_BLOCK

FUNCTION_BLOCK "ARRAY_GAV"   // FB13, SCL
TITLE = ARRAY_GAV
{ S7_Optimized_Access := 'FALSE' }
AUTHOR : hugo
FAMILY : ARFUNCT
NAME : AR_GAV
VERSION : 1.1
// this function will calculate the geometric average of a given array.
// the function needs to be called:    array_avg(adr("array"),sizeof("array"));
// because this function works with pointers its very time efficient and it needs no extra memory.
//  
// uses: SQRTN [FC112]
   VAR_INPUT
      pt : Pointer;
      _pt AT pt : Struct
         DBNr : Word;
         Adr : DWord;
      END_STRUCT;
      size : Int;
   END_VAR
   VAR_OUTPUT
      _GAV : Real;
   END_VAR
   VAR_TEMP
      i : Int;
      stop : Int;
      Adr : Int;
      DB_LENGTH : Word;
      WRITE_PROT : Bool;
      rTEST_DB : Int;
   END_VAR
BEGIN


   #_GAV := 0.0;

   (* test data block *)
   #rTEST_DB := TEST_DB(DB_NUMBER := #_pt.DBNr ,DB_LENGTH => #DB_LENGTH ,WRITE_PROT => #WRITE_PROT);
   (* End if TEST_DB <> 0 = Error *)
   IF #rTEST_DB <> 0 THEN RETURN; END_IF;
   (* End if data block to short *) 
   IF WORD_TO_INT(#DB_LENGTH)/4 < #size THEN RETURN; END_IF;
   (* calculate adress for first data *)  
   #Adr := DWORD_TO_INT(SHR(IN:=SHL(IN:=#_pt.Adr,N:=8),N:=11));

   (* code *)
   #stop := #size - 1;   //stop := SHR(size,2)-1;
   #_GAV := 1.0;
   FOR #i := 0 TO #stop DO
       IF DWORD_TO_REAL(WORD_TO_BLOCK_DB(#_pt.DBNr).DD(#Adr+#i*4)) > 0.0 THEN
           #_GAV := #_GAV * DWORD_TO_REAL(WORD_TO_BLOCK_DB(#_pt.DBNr).DD(#Adr+#i*4));
       ELSE
           #_GAV := 0.0;
           RETURN;
       END_IF;
   END_FOR;
   #_GAV := "SQRTN"(X:=#_GAV,N:=#stop+1);


   (* revision history
   hm  2. apr 2008 rev 1.0
       original version

   hm  10. mar. 2009   rev 1.1
       real constants updated to new systax using dot

   *)
END_FUNCTION_BLOCK

FUNCTION_BLOCK "ARRAY_HAV"   // FB14, SCL
TITLE = ARRAY_HAV
{ S7_Optimized_Access := 'FALSE' }
AUTHOR : hugo
FAMILY : ARFUNCT
NAME : AR_HAV
VERSION : 1.1
// this function will calculate the harmonic average of a given array.
// the function needs to be called:    array_avg(adr("array"),sizeof("array"));
// because this function works with pointers its very time efficient and it needs no extra memory.
   VAR_INPUT
      pt : Pointer;
      _pt AT pt : Struct
         DBNr : Word;
         Adr : DWord;
      END_STRUCT;
      size : Int;
   END_VAR
   VAR_OUTPUT
      _HAV : Real;
   END_VAR
   VAR_TEMP
      i : Int;
      stop : Int;
      Adr : Int;
      DB_LENGTH : Word;
      WRITE_PROT : Bool;
      rTEST_DB : Int;
   END_VAR
BEGIN


   #_HAV := 0.0;

   (* test data block *)
   #rTEST_DB := TEST_DB(DB_NUMBER := #_pt.DBNr ,DB_LENGTH => #DB_LENGTH ,WRITE_PROT => #WRITE_PROT);
   (* End if TEST_DB <> 0 = Error *)
   IF #rTEST_DB <> 0 THEN RETURN; END_IF;
   (* End if data block to short *) 
   IF WORD_TO_INT(#DB_LENGTH)/4 < #size THEN RETURN; END_IF;
   (* calculate adress for first data *)  
   #Adr := DWORD_TO_INT(SHR(IN:=SHL(IN:=#_pt.Adr,N:=8),N:=11));

   (* code *)
   #stop := #size - 1;   //stop := SHR(size,2)-1;
   FOR #i := 0 TO #stop DO
       IF DWORD_TO_REAL(WORD_TO_BLOCK_DB(#_pt.DBNr).DD(#Adr+#i*4)) <> 0.0 THEN
           #_HAV := #_HAV + 1.0/DWORD_TO_REAL(WORD_TO_BLOCK_DB(#_pt.DBNr).DD(#Adr+#i*4));
       ELSE
           #_HAV := 0.0;
           RETURN;
       END_IF;
   END_FOR;
   #_HAV := (INT_TO_REAL(#stop) + 1.0) / #_HAV;


   (* revision history
   hm  2. apr 2008 rev 1.0
       original version

   hm  10. mar. 2009   rev 1.1
       real constants updated to new systax using dot

   *)
END_FUNCTION_BLOCK

FUNCTION_BLOCK "ARRAY_MAX"   // FB15, SCL
TITLE = ARRAY_MAX
{ S7_Optimized_Access := 'FALSE' }
AUTHOR : hugo
FAMILY : ARFUNCT
NAME : AR_MAX
VERSION : 1.1
// this function will calculate the max value of a given array.
// the function needs to be called:    array_max(adr("array"),sizeof("array"));
// because this function works with pointers its very time efficient and it needs no extra memory.
   VAR_INPUT
      pt : Pointer;
      _pt AT pt : Struct
         DBNr : Word;
         Adr : DWord;
      END_STRUCT;
      size : Int;
   END_VAR
   VAR_OUTPUT
      _max : Real;
   END_VAR
   VAR_TEMP
      i : Int;
      Adr : Int;
      DB_LENGTH : Word;
      WRITE_PROT : Bool;
      rTEST_DB : Int;
   END_VAR
BEGIN


     (* Datenbaustein Testen *)
     #rTEST_DB := TEST_DB(DB_NUMBER := #_pt.DBNr // IN: WORD
                        ,DB_LENGTH => #DB_LENGTH // OUT: WORD
                        ,WRITE_PROT => #WRITE_PROT // OUT: BOOL
                        ); // INT
     (* Ende wenn Test-DB <> 0 = Fehler *)
     IF #rTEST_DB <> 0 THEN RETURN; END_IF;
     (* Ende wenn DB zu klein *) 
     IF WORD_TO_INT(#DB_LENGTH)/4 < #size THEN RETURN; END_IF;

     #Adr := DWORD_TO_INT(SHR(IN:=SHL(IN:=#_pt.Adr,N:=8),N:=11));

     (* Berechnung *)
     #_max := DWORD_TO_REAL(WORD_TO_BLOCK_DB(#_pt.DBNr).DD(#Adr+0));
     FOR #i := 1 TO #size-1 DO
         IF DWORD_TO_REAL(WORD_TO_BLOCK_DB(#_pt.DBNr).DD(#Adr+#i*4)) > #_max THEN 
             #_max := DWORD_TO_REAL(WORD_TO_BLOCK_DB(#_pt.DBNr).DD(#Adr+#i*4)); 
         END_IF;
     END_FOR;

   (* revision history
   hm  2. oct 2006     rev 1.0
       original version

   hm  16. mar. 2008   rev 1.1
       changed input size to uint
   *)
END_FUNCTION_BLOCK

FUNCTION_BLOCK "ARRAY_MIN"   // FB16, SCL
TITLE = ARRAY_MIN
{ S7_Optimized_Access := 'FALSE' }
AUTHOR : hugo
FAMILY : ARFUNCT
NAME : AR_MIN
VERSION : 1.1
// this function will calculate the min value of a given array.
// the function needs to be called:    array_min(adr("array"),sizeof("array"));
// because this function works with pointers its very time efficient and it needs no extra memory.
   VAR_INPUT
      pt : Pointer;
      _pt AT pt : Struct
         DBNr : Word;
         Adr : DWord;
      END_STRUCT;
      size : Int;
   END_VAR
   VAR_OUTPUT
      _min : Real;
   END_VAR
   VAR_TEMP
      i : Int;
      Adr : Int;
      DB_LENGTH : Word;
      WRITE_PROT : Bool;
      rTEST_DB : Int;
   END_VAR
BEGIN


     (* Datenbaustein Testen *)
     #rTEST_DB := TEST_DB(DB_NUMBER := #_pt.DBNr // IN: WORD
                        ,DB_LENGTH => #DB_LENGTH // OUT: WORD
                        ,WRITE_PROT => #WRITE_PROT // OUT: BOOL
                        ); // INT
     (* Ende wenn Test-DB <> 0 = Fehler *)
     IF #rTEST_DB <> 0 THEN RETURN; END_IF;
     (* Ende wenn DB zu klein *) 
     IF WORD_TO_INT(#DB_LENGTH)/4 < #size THEN RETURN; END_IF;

     #Adr := DWORD_TO_INT(SHR(IN:=SHL(IN:=#_pt.Adr,N:=8),N:=11));

     (* Berechnung *)
     #_min := DWORD_TO_REAL(WORD_TO_BLOCK_DB(#_pt.DBNr).DD(#Adr+0));
     FOR #i := 1 TO #size-1 DO
         IF DWORD_TO_REAL(WORD_TO_BLOCK_DB(#_pt.DBNr).DD(#Adr+#i*4)) < #_min THEN 
             #_min := DWORD_TO_REAL(WORD_TO_BLOCK_DB(#_pt.DBNr).DD(#Adr+#i*4)); 
         END_IF;
     END_FOR;

   (* revision history
   hm      2. oct. 2006
       original version

   hm      16. mar. 2008
       changed type of input size to uint

   *)
END_FUNCTION_BLOCK

FUNCTION_BLOCK "ARRAY_SDV"   // FB17, SCL
TITLE = ARRAY_SDV
{ S7_Optimized_Access := 'FALSE' }
AUTHOR : hugo
FAMILY : ARFUNCT
NAME : AR_SDV
VERSION : 1.1
// this function will calculate the standard deviation of a given array.
// the function needs to be called:    array_sdv(adr("array"),sizeof("array"));
// because this function works with pointers its very time efficient and it needs no extra memory.
   VAR_INPUT
      pt : Pointer;
      _pt AT pt : Struct
         DBNr : Word;
         Adr : DWord;
      END_STRUCT;
      size : Int;
   END_VAR
   VAR_OUTPUT
      sdv : Real;
   END_VAR
   VAR_TEMP
      i : Int;
      stop : Int;
      avg : Real;
      _var : Real;
      Adr : Int;
      DB_LENGTH : Word;
      WRITE_PROT : Bool;
      rTEST_DB : Int;
   END_VAR
BEGIN


